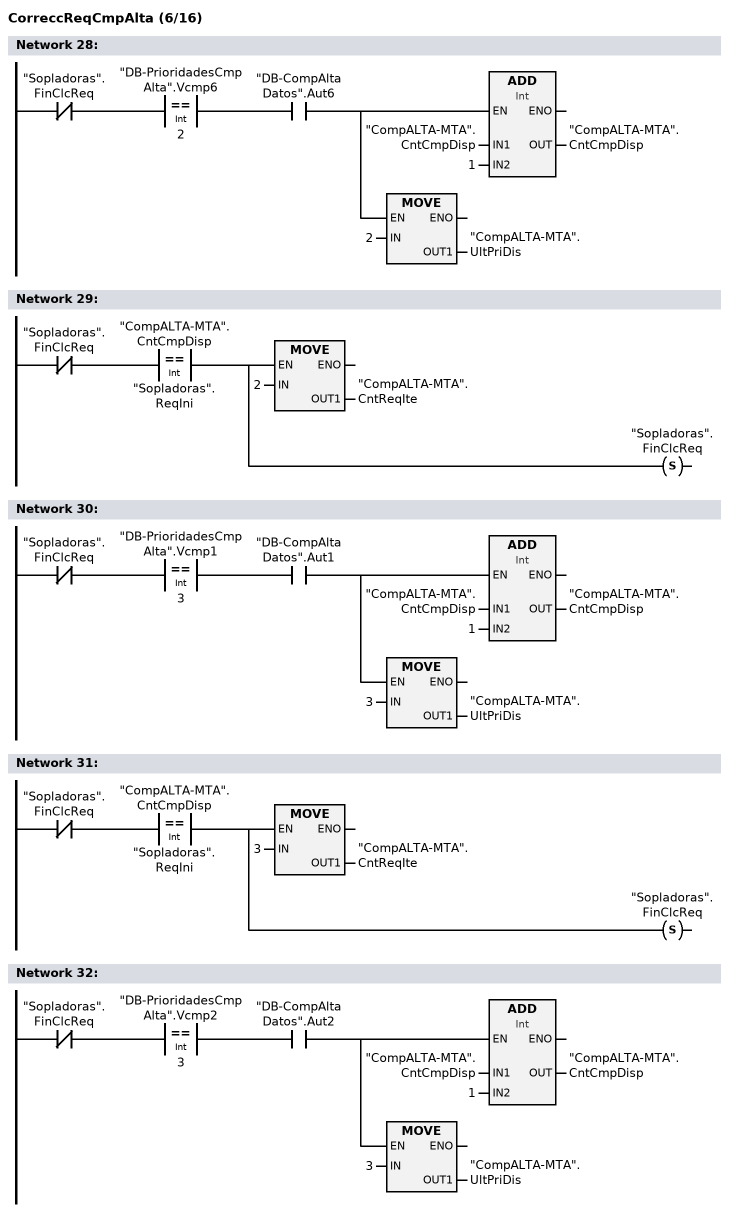
   RUNG wire#powerrail
      I_Contact( "Sopladoras".FinClcReq )
      { S7_Templates := "SrcType := Int" } EQ_Contact(in1 := "DB-PrioridadesCmpAlta".Vcmp6, in2 := 2)
      Contact( "DB-CompAltaDatos".Aut6 )
      wire#w1
      { S7_Templates := "SrcType := Int"; S7_GenerateENO := "TRUE" } Add(in1 := "CompALTA-MTA".CntCmpDisp, in2 := 1, out => "CompALTA-MTA".CntCmpDisp)
   END_RUNG
   RUNG wire#w1
      { S7_GenerateENO := "TRUE" } Move(in := 2, out1 => "CompALTA-MTA".UltPriDis)
   END_RUNG
   // the same network as SCL:
   IF NOT "Sopladoras".FinClcReq AND ("DB-PrioridadesCmpAlta".Vcmp6 = 2) AND "DB-CompAltaDatos".Aut6 THEN
       "CompALTA-MTA".CntCmpDisp := "CompALTA-MTA".CntCmpDisp + 1;
       "CompALTA-MTA".UltPriDis := 2;
   END_IF;
END_REGION

REGION Network 29
   RUNG wire#powerrail
      I_Contact( "Sopladoras".FinClcReq )
      { S7_Templates := "SrcType := Int" } EQ_Contact(in1 := "CompALTA-MTA".CntCmpDisp, in2 := "Sopladoras".ReqIni)
      wire#w1
      { S7_GenerateENO := "TRUE" } Move(in := 2, out1 => "CompALTA-MTA".CntReqIte)
   END_RUNG
   RUNG wire#w1
      S_Coil( "Sopladoras".FinClcReq )
   END_RUNG
   // the same network as SCL:
   IF NOT "Sopladoras".FinClcReq AND ("CompALTA-MTA".CntCmpDisp = "Sopladoras".ReqIni) THEN
       "CompALTA-MTA".CntReqIte := 2;
       "Sopladoras".FinClcReq := TRUE;
   END_IF;
END_REGION

REGION Network 30
   IF NOT "Sopladoras".FinClcReq AND ("DB-PrioridadesCmpAlta".Vcmp1 = 3) AND "DB-CompAltaDatos".Aut1 THEN
       "CompALTA-MTA".CntCmpDisp := "CompALTA-MTA".CntCmpDisp + 1;
       "CompALTA-MTA".UltPriDis := 3;
   END_IF;
END_REGION

REGION Network 31
   IF NOT "Sopladoras".FinClcReq AND ("CompALTA-MTA".CntCmpDisp = "Sopladoras".ReqIni) THEN
       "CompALTA-MTA".CntReqIte := 3;
       "Sopladoras".FinClcReq := TRUE;
   END_IF;
END_REGION

REGION Network 32
   IF NOT "Sopladoras".FinClcReq AND ("DB-PrioridadesCmpAlta".Vcmp2 = 3) AND "DB-CompAltaDatos".Aut2 THEN
       "CompALTA-MTA".CntCmpDisp := "CompALTA-MTA".CntCmpDisp + 1;
       "CompALTA-MTA".UltPriDis := 3;
   END_IF;
END_REGION

REGION Network 33
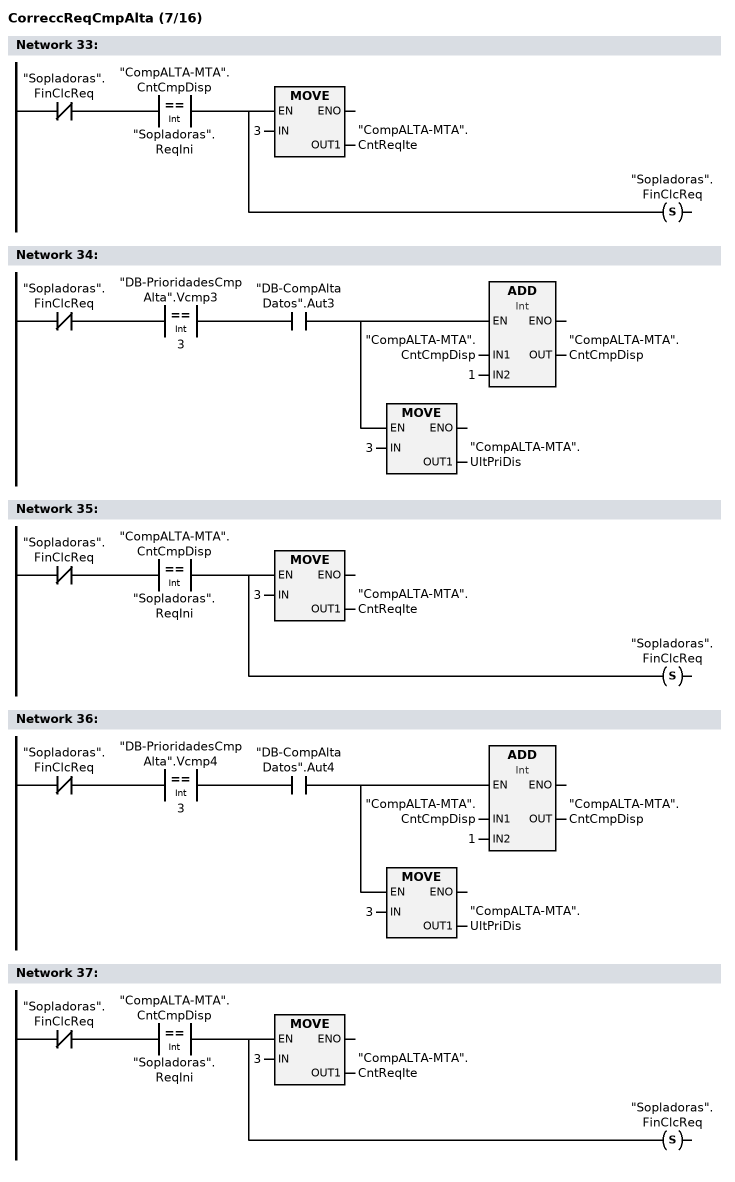
   IF NOT "Sopladoras".FinClcReq AND ("CompALTA-MTA".CntCmpDisp = "Sopladoras".ReqIni) THEN
       "CompALTA-MTA".CntReqIte := 3;
       "Sopladoras".FinClcReq := TRUE;
   END_IF;
END_REGION

REGION Network 34
   IF NOT "Sopladoras".FinClcReq AND ("DB-PrioridadesCmpAlta".Vcmp3 = 3) AND "DB-CompAltaDatos".Aut3 THEN
       "CompALTA-MTA".CntCmpDisp := "CompALTA-MTA".CntCmpDisp + 1;
       "CompALTA-MTA".UltPriDis := 3;
   END_IF;
END_REGION

REGION Network 35
   IF NOT "Sopladoras".FinClcReq AND ("CompALTA-MTA".CntCmpDisp = "Sopladoras".ReqIni) THEN
       "CompALTA-MTA".CntReqIte := 3;
       "Sopladoras".FinClcReq := TRUE;
   END_IF;
END_REGION

REGION Network 36
   IF NOT "Sopladoras".FinClcReq AND ("DB-PrioridadesCmpAlta".Vcmp4 = 3) AND "DB-CompAltaDatos".Aut4 THEN
       "CompALTA-MTA".CntCmpDisp := "CompALTA-MTA".CntCmpDisp + 1;
       "CompALTA-MTA".UltPriDis := 3;
   END_IF;
END_REGION

REGION Network 37
   IF NOT "Sopladoras".FinClcReq AND ("CompALTA-MTA".CntCmpDisp = "Sopladoras".ReqIni) THEN
       "CompALTA-MTA".CntReqIte := 3;
       "Sopladoras".FinClcReq := TRUE;
   END_IF;
END_REGION

REGION Network 38
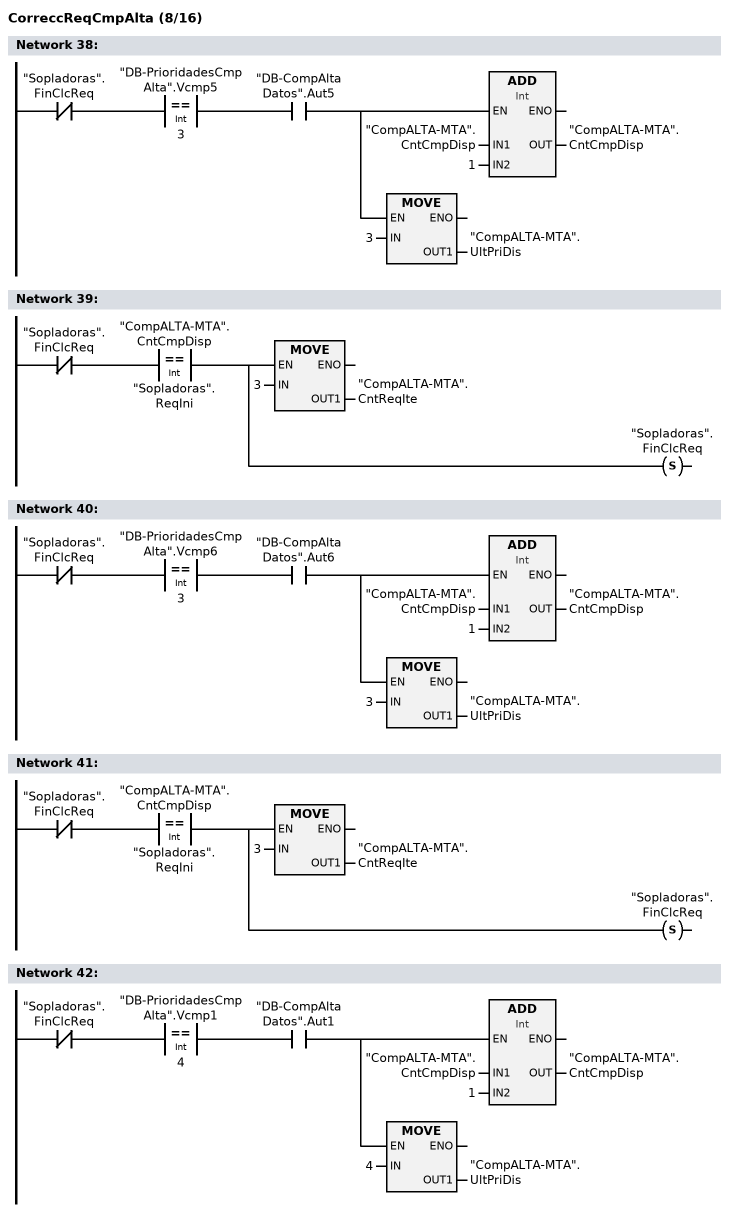
   IF NOT "Sopladoras".FinClcReq AND ("DB-PrioridadesCmpAlta".Vcmp5 = 3) AND "DB-CompAltaDatos".Aut5 THEN
       "CompALTA-MTA".CntCmpDisp := "CompALTA-MTA".CntCmpDisp + 1;
       "CompALTA-MTA".UltPriDis := 3;
   END_IF;
END_REGION

REGION Network 39
   IF NOT "Sopladoras".FinClcReq AND ("CompALTA-MTA".CntCmpDisp = "Sopladoras".ReqIni) THEN
       "CompALTA-MTA".CntReqIte := 3;
       "Sopladoras".FinClcReq := TRUE;
   END_IF;
END_REGION

REGION Network 40
   RUNG wire#powerrail
      I_Contact( "Sopladoras".FinClcReq )
      { S7_Templates := "SrcType := Int" } EQ_Contact(in1 := "DB-PrioridadesCmpAlta".Vcmp6, in2 := 3)
      Contact( "DB-CompAltaDatos".Aut6 )
      wire#w1
      { S7_Templates := "SrcType := Int"; S7_GenerateENO := "TRUE" } Add(in1 := "CompALTA-MTA".CntCmpDisp, in2 := 1, out => "CompALTA-MTA".CntCmpDisp)
   END_RUNG
   RUNG wire#w1
      { S7_GenerateENO := "TRUE" } Move(in := 3, out1 => "CompALTA-MTA".UltPriDis)
   END_RUNG
   // the same network as SCL:
   IF NOT "Sopladoras".FinClcReq AND ("DB-PrioridadesCmpAlta".Vcmp6 = 3) AND "DB-CompAltaDatos".Aut6 THEN
       "CompALTA-MTA".CntCmpDisp := "CompALTA-MTA".CntCmpDisp + 1;
       "CompALTA-MTA".UltPriDis := 3;
   END_IF;
END_REGION

REGION Network 41
   RUNG wire#powerrail
      I_Contact( "Sopladoras".FinClcReq )
      { S7_Templates := "SrcType := Int" } EQ_Contact(in1 := "CompALTA-MTA".CntCmpDisp, in2 := "Sopladoras".ReqIni)
      wire#w1
      { S7_GenerateENO := "TRUE" } Move(in := 3, out1 => "CompALTA-MTA".CntReqIte)
   END_RUNG
   RUNG wire#w1
      S_Coil( "Sopladoras".FinClcReq )
   END_RUNG
   // the same network as SCL:
   IF NOT "Sopladoras".FinClcReq AND ("CompALTA-MTA".CntCmpDisp = "Sopladoras".ReqIni) THEN
       "CompALTA-MTA".CntReqIte := 3;
       "Sopladoras".FinClcReq := TRUE;
   END_IF;
END_REGION

REGION Network 42
   IF NOT "Sopladoras".FinClcReq AND ("DB-PrioridadesCmpAlta".Vcmp1 = 4) AND "DB-CompAltaDatos".Aut1 THEN
       "CompALTA-MTA".CntCmpDisp := "CompALTA-MTA".CntCmpDisp + 1;
       "CompALTA-MTA".UltPriDis := 4;
   END_IF;
END_REGION

REGION Network 43
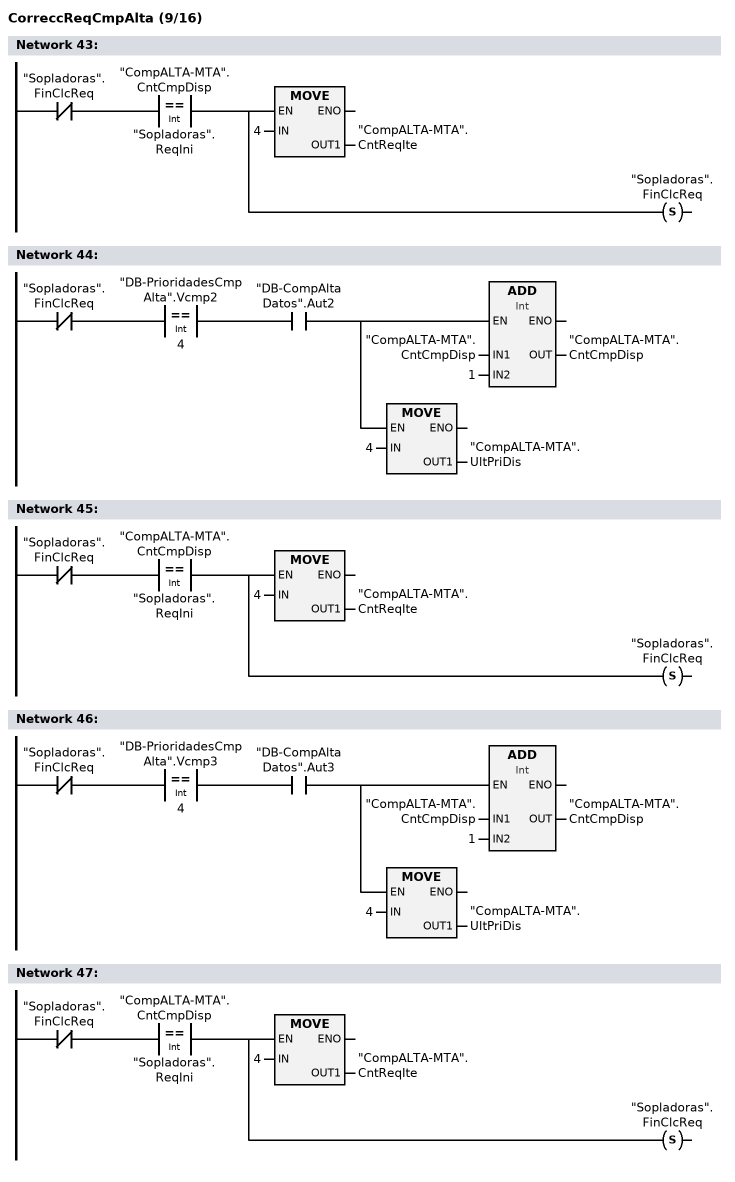
   IF NOT "Sopladoras".FinClcReq AND ("CompALTA-MTA".CntCmpDisp = "Sopladoras".ReqIni) THEN
       "CompALTA-MTA".CntReqIte := 4;
       "Sopladoras".FinClcReq := TRUE;
   END_IF;
END_REGION

REGION Network 44
   IF NOT "Sopladoras".FinClcReq AND ("DB-PrioridadesCmpAlta".Vcmp2 = 4) AND "DB-CompAltaDatos".Aut2 THEN
       "CompALTA-MTA".CntCmpDisp := "CompALTA-MTA".CntCmpDisp + 1;
       "CompALTA-MTA".UltPriDis := 4;
   END_IF;
END_REGION

REGION Network 45
   IF NOT "Sopladoras".FinClcReq AND ("CompALTA-MTA".CntCmpDisp = "Sopladoras".ReqIni) THEN
       "CompALTA-MTA".CntReqIte := 4;
       "Sopladoras".FinClcReq := TRUE;
   END_IF;
END_REGION

REGION Network 46
   IF NOT "Sopladoras".FinClcReq AND ("DB-PrioridadesCmpAlta".Vcmp3 = 4) AND "DB-CompAltaDatos".Aut3 THEN
       "CompALTA-MTA".CntCmpDisp := "CompALTA-MTA".CntCmpDisp + 1;
       "CompALTA-MTA".UltPriDis := 4;
   END_IF;
END_REGION

REGION Network 47
   IF NOT "Sopladoras".FinClcReq AND ("CompALTA-MTA".CntCmpDisp = "Sopladoras".ReqIni) THEN
       "CompALTA-MTA".CntReqIte := 4;
       "Sopladoras".FinClcReq := TRUE;
   END_IF;
END_REGION

REGION Network 48
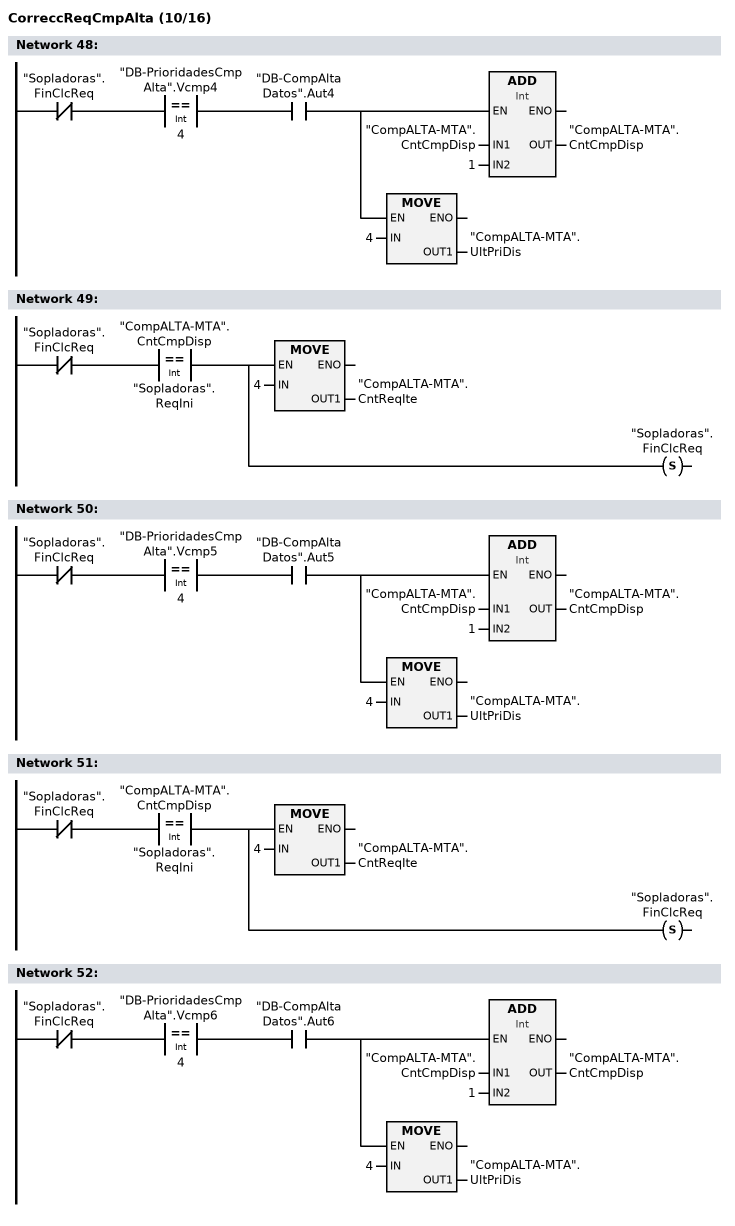
   IF NOT "Sopladoras".FinClcReq AND ("DB-PrioridadesCmpAlta".Vcmp4 = 4) AND "DB-CompAltaDatos".Aut4 THEN
       "CompALTA-MTA".CntCmpDisp := "CompALTA-MTA".CntCmpDisp + 1;
       "CompALTA-MTA".UltPriDis := 4;
   END_IF;
END_REGION

REGION Network 49
   IF NOT "Sopladoras".FinClcReq AND ("CompALTA-MTA".CntCmpDisp = "Sopladoras".ReqIni) THEN
       "CompALTA-MTA".CntReqIte := 4;
       "Sopladoras".FinClcReq := TRUE;
   END_IF;
END_REGION

REGION Network 50
   IF NOT "Sopladoras".FinClcReq AND ("DB-PrioridadesCmpAlta".Vcmp5 = 4) AND "DB-CompAltaDatos".Aut5 THEN
       "CompALTA-MTA".CntCmpDisp := "CompALTA-MTA".CntCmpDisp + 1;
       "CompALTA-MTA".UltPriDis := 4;
   END_IF;
END_REGION

REGION Network 51
   IF NOT "Sopladoras".FinClcReq AND ("CompALTA-MTA".CntCmpDisp = "Sopladoras".ReqIni) THEN
       "CompALTA-MTA".CntReqIte := 4;
       "Sopladoras".FinClcReq := TRUE;
   END_IF;
END_REGION

REGION Network 52
   RUNG wire#powerrail
      I_Contact( "Sopladoras".FinClcReq )
      { S7_Templates := "SrcType := Int" } EQ_Contact(in1 := "DB-PrioridadesCmpAlta".Vcmp6, in2 := 4)
      Contact( "DB-CompAltaDatos".Aut6 )
      wire#w1
      { S7_Templates := "SrcType := Int"; S7_GenerateENO := "TRUE" } Add(in1 := "CompALTA-MTA".CntCmpDisp, in2 := 1, out => "CompALTA-MTA".CntCmpDisp)
   END_RUNG
   RUNG wire#w1
      { S7_GenerateENO := "TRUE" } Move(in := 4, out1 => "CompALTA-MTA".UltPriDis)
   END_RUNG
   // the same network as SCL:
   IF NOT "Sopladoras".FinClcReq AND ("DB-PrioridadesCmpAlta".Vcmp6 = 4) AND "DB-CompAltaDatos".Aut6 THEN
       "CompALTA-MTA".CntCmpDisp := "CompALTA-MTA".CntCmpDisp + 1;
       "CompALTA-MTA".UltPriDis := 4;
   END_IF;
END_REGION

REGION Network 53
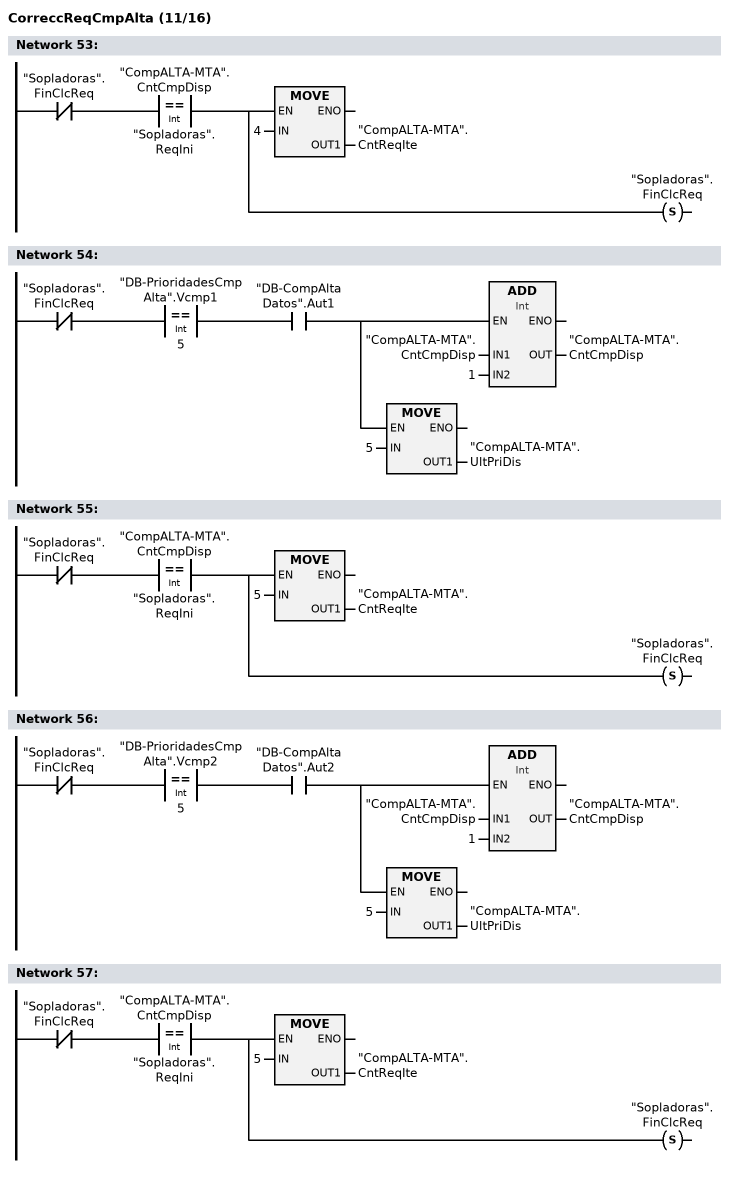
   RUNG wire#powerrail
      I_Contact( "Sopladoras".FinClcReq )
      { S7_Templates := "SrcType := Int" } EQ_Contact(in1 := "CompALTA-MTA".CntCmpDisp, in2 := "Sopladoras".ReqIni)
      wire#w1
      { S7_GenerateENO := "TRUE" } Move(in := 4, out1 => "CompALTA-MTA".CntReqIte)
   END_RUNG
   RUNG wire#w1
      S_Coil( "Sopladoras".FinClcReq )
   END_RUNG
   // the same network as SCL:
   IF NOT "Sopladoras".FinClcReq AND ("CompALTA-MTA".CntCmpDisp = "Sopladoras".ReqIni) THEN
       "CompALTA-MTA".CntReqIte := 4;
       "Sopladoras".FinClcReq := TRUE;
   END_IF;
END_REGION

REGION Network 54
   IF NOT "Sopladoras".FinClcReq AND ("DB-PrioridadesCmpAlta".Vcmp1 = 5) AND "DB-CompAltaDatos".Aut1 THEN
       "CompALTA-MTA".CntCmpDisp := "CompALTA-MTA".CntCmpDisp + 1;
       "CompALTA-MTA".UltPriDis := 5;
   END_IF;
END_REGION

REGION Network 55
   IF NOT "Sopladoras".FinClcReq AND ("CompALTA-MTA".CntCmpDisp = "Sopladoras".ReqIni) THEN
       "CompALTA-MTA".CntReqIte := 5;
       "Sopladoras".FinClcReq := TRUE;
   END_IF;
END_REGION

REGION Network 56
   IF NOT "Sopladoras".FinClcReq AND ("DB-PrioridadesCmpAlta".Vcmp2 = 5) AND "DB-CompAltaDatos".Aut2 THEN
       "CompALTA-MTA".CntCmpDisp := "CompALTA-MTA".CntCmpDisp + 1;
       "CompALTA-MTA".UltPriDis := 5;
   END_IF;
END_REGION

REGION Network 57
   IF NOT "Sopladoras".FinClcReq AND ("CompALTA-MTA".CntCmpDisp = "Sopladoras".ReqIni) THEN
       "CompALTA-MTA".CntReqIte := 5;
       "Sopladoras".FinClcReq := TRUE;
   END_IF;
END_REGION

REGION Network 58
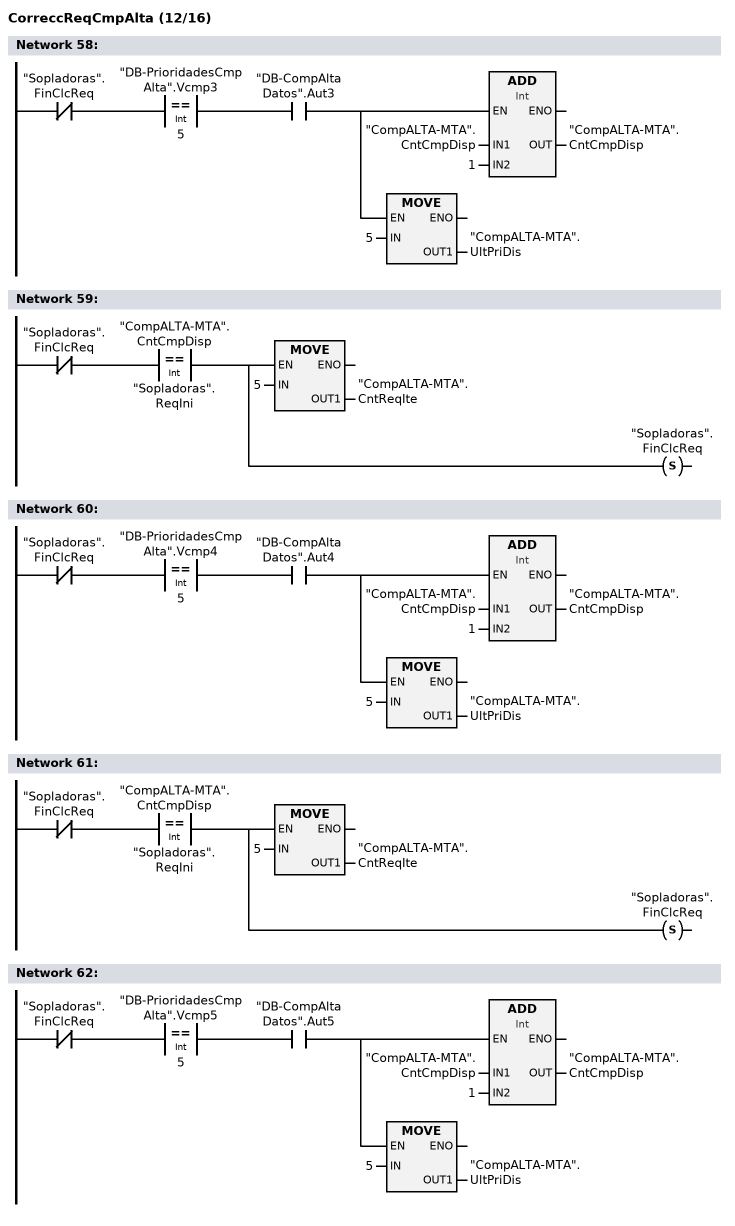
   IF NOT "Sopladoras".FinClcReq AND ("DB-PrioridadesCmpAlta".Vcmp3 = 5) AND "DB-CompAltaDatos".Aut3 THEN
       "CompALTA-MTA".CntCmpDisp := "CompALTA-MTA".CntCmpDisp + 1;
       "CompALTA-MTA".UltPriDis := 5;
   END_IF;
END_REGION

REGION Network 59
   IF NOT "Sopladoras".FinClcReq AND ("CompALTA-MTA".CntCmpDisp = "Sopladoras".ReqIni) THEN
       "CompALTA-MTA".CntReqIte := 5;
       "Sopladoras".FinClcReq := TRUE;
   END_IF;
END_REGION

REGION Network 60
   IF NOT "Sopladoras".FinClcReq AND ("DB-PrioridadesCmpAlta".Vcmp4 = 5) AND "DB-CompAltaDatos".Aut4 THEN
       "CompALTA-MTA".CntCmpDisp := "CompALTA-MTA".CntCmpDisp + 1;
       "CompALTA-MTA".UltPriDis := 5;
   END_IF;
END_REGION

REGION Network 61
   IF NOT "Sopladoras".FinClcReq AND ("CompALTA-MTA".CntCmpDisp = "Sopladoras".ReqIni) THEN
       "CompALTA-MTA".CntReqIte := 5;
       "Sopladoras".FinClcReq := TRUE;
   END_IF;
END_REGION

REGION Network 62
   IF NOT "Sopladoras".FinClcReq AND ("DB-PrioridadesCmpAlta".Vcmp5 = 5) AND "DB-CompAltaDatos".Aut5 THEN
       "CompALTA-MTA".CntCmpDisp := "CompALTA-MTA".CntCmpDisp + 1;
       "CompALTA-MTA".UltPriDis := 5;
   END_IF;
END_REGION

REGION Network 63
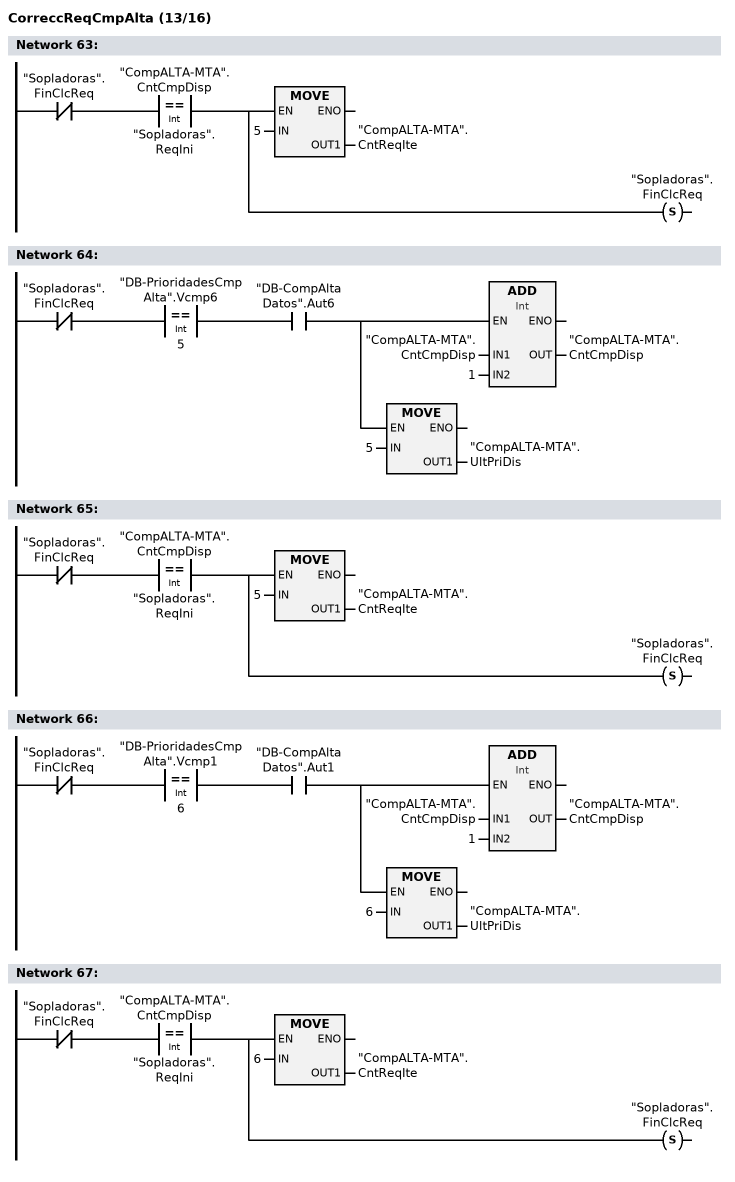
   IF NOT "Sopladoras".FinClcReq AND ("CompALTA-MTA".CntCmpDisp = "Sopladoras".ReqIni) THEN
       "CompALTA-MTA".CntReqIte := 5;
       "Sopladoras".FinClcReq := TRUE;
   END_IF;
END_REGION

REGION Network 64
   RUNG wire#powerrail
      I_Contact( "Sopladoras".FinClcReq )
      { S7_Templates := "SrcType := Int" } EQ_Contact(in1 := "DB-PrioridadesCmpAlta".Vcmp6, in2 := 5)
      Contact( "DB-CompAltaDatos".Aut6 )
      wire#w1
      { S7_Templates := "SrcType := Int"; S7_GenerateENO := "TRUE" } Add(in1 := "CompALTA-MTA".CntCmpDisp, in2 := 1, out => "CompALTA-MTA".CntCmpDisp)
   END_RUNG
   RUNG wire#w1
      { S7_GenerateENO := "TRUE" } Move(in := 5, out1 => "CompALTA-MTA".UltPriDis)
   END_RUNG
   // the same network as SCL:
   IF NOT "Sopladoras".FinClcReq AND ("DB-PrioridadesCmpAlta".Vcmp6 = 5) AND "DB-CompAltaDatos".Aut6 THEN
       "CompALTA-MTA".CntCmpDisp := "CompALTA-MTA".CntCmpDisp + 1;
       "CompALTA-MTA".UltPriDis := 5;
   END_IF;
END_REGION

REGION Network 65
   RUNG wire#powerrail
      I_Contact( "Sopladoras".FinClcReq )
      { S7_Templates := "SrcType := Int" } EQ_Contact(in1 := "CompALTA-MTA".CntCmpDisp, in2 := "Sopladoras".ReqIni)
      wire#w1
      { S7_GenerateENO := "TRUE" } Move(in := 5, out1 => "CompALTA-MTA".CntReqIte)
   END_RUNG
   RUNG wire#w1
      S_Coil( "Sopladoras".FinClcReq )
   END_RUNG
   // the same network as SCL:
   IF NOT "Sopladoras".FinClcReq AND ("CompALTA-MTA".CntCmpDisp = "Sopladoras".ReqIni) THEN
       "CompALTA-MTA".CntReqIte := 5;
       "Sopladoras".FinClcReq := TRUE;
   END_IF;
END_REGION

REGION Network 66
   RUNG wire#powerrail
      I_Contact( "Sopladoras".FinClcReq )
      { S7_Templates := "SrcType := Int" } EQ_Contact(in1 := "DB-PrioridadesCmpAlta".Vcmp1, in2 := 6)
      Contact( "DB-CompAltaDatos".Aut1 )
      wire#w1
      { S7_Templates := "SrcType := Int"; S7_GenerateENO := "TRUE" } Add(in1 := "CompALTA-MTA".CntCmpDisp, in2 := 1, out => "CompALTA-MTA".CntCmpDisp)
   END_RUNG
   RUNG wire#w1
      { S7_GenerateENO := "TRUE" } Move(in := 6, out1 => "CompALTA-MTA".UltPriDis)
   END_RUNG
   // the same network as SCL:
   IF NOT "Sopladoras".FinClcReq AND ("DB-PrioridadesCmpAlta".Vcmp1 = 6) AND "DB-CompAltaDatos".Aut1 THEN
       "CompALTA-MTA".CntCmpDisp := "CompALTA-MTA".CntCmpDisp + 1;
       "CompALTA-MTA".UltPriDis := 6;
   END_IF;
END_REGION

REGION Network 67
   RUNG wire#powerrail
      I_Contact( "Sopladoras".FinClcReq )
      { S7_Templates := "SrcType := Int" } EQ_Contact(in1 := "CompALTA-MTA".CntCmpDisp, in2 := "Sopladoras".ReqIni)
      wire#w1
      { S7_GenerateENO := "TRUE" } Move(in := 6, out1 => "CompALTA-MTA".CntReqIte)
   END_RUNG
   RUNG wire#w1
      S_Coil( "Sopladoras".FinClcReq )
   END_RUNG
   // the same network as SCL:
   IF NOT "Sopladoras".FinClcReq AND ("CompALTA-MTA".CntCmpDisp = "Sopladoras".ReqIni) THEN
       "CompALTA-MTA".CntReqIte := 6;
       "Sopladoras".FinClcReq := TRUE;
   END_IF;
END_REGION

REGION Network 68
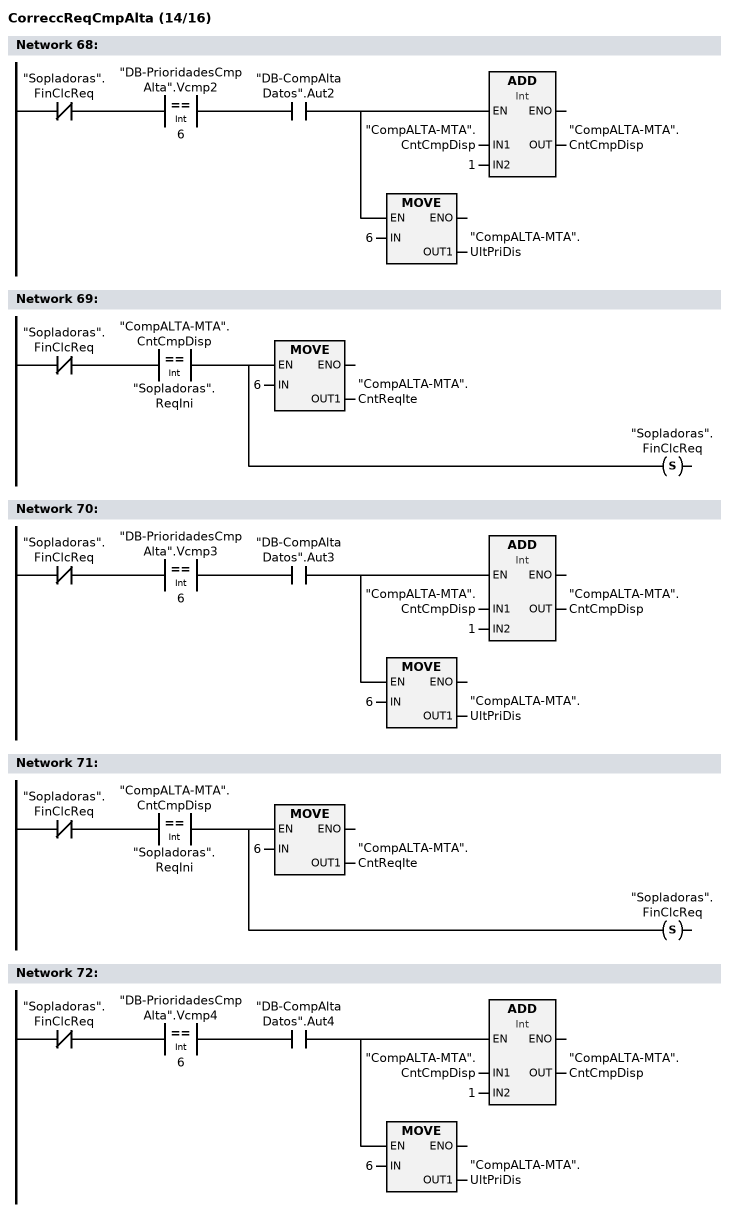
   RUNG wire#powerrail
      I_Contact( "Sopladoras".FinClcReq )
      { S7_Templates := "SrcType := Int" } EQ_Contact(in1 := "DB-PrioridadesCmpAlta".Vcmp2, in2 := 6)
      Contact( "DB-CompAltaDatos".Aut2 )
      wire#w1
      { S7_Templates := "SrcType := Int"; S7_GenerateENO := "TRUE" } Add(in1 := "CompALTA-MTA".CntCmpDisp, in2 := 1, out => "CompALTA-MTA".CntCmpDisp)
   END_RUNG
   RUNG wire#w1
      { S7_GenerateENO := "TRUE" } Move(in := 6, out1 => "CompALTA-MTA".UltPriDis)
   END_RUNG
   // the same network as SCL:
   IF NOT "Sopladoras".FinClcReq AND ("DB-PrioridadesCmpAlta".Vcmp2 = 6) AND "DB-CompAltaDatos".Aut2 THEN
       "CompALTA-MTA".CntCmpDisp := "CompALTA-MTA".CntCmpDisp + 1;
       "CompALTA-MTA".UltPriDis := 6;
   END_IF;
END_REGION

REGION Network 69
   RUNG wire#powerrail
      I_Contact( "Sopladoras".FinClcReq )
      { S7_Templates := "SrcType := Int" } EQ_Contact(in1 := "CompALTA-MTA".CntCmpDisp, in2 := "Sopladoras".ReqIni)
      wire#w1
      { S7_GenerateENO := "TRUE" } Move(in := 6, out1 => "CompALTA-MTA".CntReqIte)
   END_RUNG
   RUNG wire#w1
      S_Coil( "Sopladoras".FinClcReq )
   END_RUNG
   // the same network as SCL:
   IF NOT "Sopladoras".FinClcReq AND ("CompALTA-MTA".CntCmpDisp = "Sopladoras".ReqIni) THEN
       "CompALTA-MTA".CntReqIte := 6;
       "Sopladoras".FinClcReq := TRUE;
   END_IF;
END_REGION

REGION Network 70
   RUNG wire#powerrail
      I_Contact( "Sopladoras".FinClcReq )
      { S7_Templates := "SrcType := Int" } EQ_Contact(in1 := "DB-PrioridadesCmpAlta".Vcmp3, in2 := 6)
      Contact( "DB-CompAltaDatos".Aut3 )
      wire#w1
      { S7_Templates := "SrcType := Int"; S7_GenerateENO := "TRUE" } Add(in1 := "CompALTA-MTA".CntCmpDisp, in2 := 1, out => "CompALTA-MTA".CntCmpDisp)
   END_RUNG
   RUNG wire#w1
      { S7_GenerateENO := "TRUE" } Move(in := 6, out1 => "CompALTA-MTA".UltPriDis)
   END_RUNG
   // the same network as SCL:
   IF NOT "Sopladoras".FinClcReq AND ("DB-PrioridadesCmpAlta".Vcmp3 = 6) AND "DB-CompAltaDatos".Aut3 THEN
       "CompALTA-MTA".CntCmpDisp := "CompALTA-MTA".CntCmpDisp + 1;
       "CompALTA-MTA".UltPriDis := 6;
   END_IF;
END_REGION

REGION Network 71
   RUNG wire#powerrail
      I_Contact( "Sopladoras".FinClcReq )
      { S7_Templates := "SrcType := Int" } EQ_Contact(in1 := "CompALTA-MTA".CntCmpDisp, in2 := "Sopladoras".ReqIni)
      wire#w1
      { S7_GenerateENO := "TRUE" } Move(in := 6, out1 => "CompALTA-MTA".CntReqIte)
   END_RUNG
   RUNG wire#w1
      S_Coil( "Sopladoras".FinClcReq )
   END_RUNG
   // the same network as SCL:
   IF NOT "Sopladoras".FinClcReq AND ("CompALTA-MTA".CntCmpDisp = "Sopladoras".ReqIni) THEN
       "CompALTA-MTA".CntReqIte := 6;
       "Sopladoras".FinClcReq := TRUE;
   END_IF;
END_REGION

REGION Network 72
   RUNG wire#powerrail
      I_Contact( "Sopladoras".FinClcReq )
      { S7_Templates := "SrcType := Int" } EQ_Contact(in1 := "DB-PrioridadesCmpAlta".Vcmp4, in2 := 6)
      Contact( "DB-CompAltaDatos".Aut4 )
      wire#w1
      { S7_Templates := "SrcType := Int"; S7_GenerateENO := "TRUE" } Add(in1 := "CompALTA-MTA".CntCmpDisp, in2 := 1, out => "CompALTA-MTA".CntCmpDisp)
   END_RUNG
   RUNG wire#w1
      { S7_GenerateENO := "TRUE" } Move(in := 6, out1 => "CompALTA-MTA".UltPriDis)
   END_RUNG
   // the same network as SCL:
   IF NOT "Sopladoras".FinClcReq AND ("DB-PrioridadesCmpAlta".Vcmp4 = 6) AND "DB-CompAltaDatos".Aut4 THEN
       "CompALTA-MTA".CntCmpDisp := "CompALTA-MTA".CntCmpDisp + 1;
       "CompALTA-MTA".UltPriDis := 6;
   END_IF;
END_REGION

REGION Network 73